VAR_GLOBAL   // PLC tag table "RIO_6"
   "Tank 6P GTT Isolation Valve Feedback - Opened" AT %I60.0 : Bool;   // CV422-6P
   "Tank 6P GTT Isolation Valve Feedback - Closed" AT %I60.1 : Bool;   // CV422-6P
   "Tank 6P Tank Vent Valve 1 Feedback - Opened" AT %I60.2 : Bool;   // CV441-6PA
   "Tank 6P Tank Vent Valve 1 Feedback - Closed" AT %I60.3 : Bool;   // CV441-6PA
   "Tank 6P Tank Vent Valve 2 Feedback - Opened" AT %I60.4 : Bool;   // CV441-6PB
   "Tank 6P Tank Vent Valve 2 Feedback - Closed" AT %I60.5 : Bool;   // CV441-6PB
   "RIO6_SPR_DI_60_6" AT %I60.6 : Bool;   // Spare input
   "RIO6_SPR_DI_60_7" AT %I60.7 : Bool;   // Spare input
   "Tank 6S GTT Isolation Valve Feedback - Opened" AT %I63.0 : Bool;   // CV421-6S
   "Tank 6S GTT Isolation Valve Feedback - Closed" AT %I63.1 : Bool;   // CV421-6S
   "Tank 6S Tank Vent Valve 1 Feedback - Opened" AT %I63.2 : Bool;   // CV440-6SA
   "Tank 6S Tank Vent Valve 1 Feedback - Closed" AT %I63.3 : Bool;   // CV440-6SA
   "Tank 6S Tank Vent Valve 2 Feedback - Opened" AT %I63.4 : Bool;   // CV440-6SB
   "Tank 6S Tank Vent Valve 2 Feedback - Closed" AT %I63.5 : Bool;   // CV440-6SB
   "RIO6_SPR_DI_63_6" AT %I63.6 : Bool;   // Spare input
   "RIO6_SPR_DI_63_7" AT %I63.7 : Bool;   // Spare input
   "Tank 6P BWT Level High High Switch" AT %I66.0 : Bool;   // LS425-6P
   "RIO6 Tanks Pressure Switch Hi Hi" AT %I66.1 : Bool;   // PS436-6P/6S
   "Tank 6S BWT Level High High Switch" AT %I66.2 : Bool;   // LS422-6S
   "RIO6_SPR_DI_66_3" AT %I66.3 : Bool;   // Spare input
   "RIO6_SPR_DI_66_4" AT %I66.4 : Bool;   // Spare input
   "RIO6_SPR_DI_66_5" AT %I66.5 : Bool;   // Spare input
   "RIO6_SPR_DI_66_6" AT %I66.6 : Bool;   // Spare input
   "RIO6_SPR_DI_66_7" AT %I66.7 : Bool;   // Spare input
   "Tank 6P USD Flow Meter" AT %IW332 : Int;   // FIT418-6P
   "Tank 6P MBG Flow Meter" AT %IW334 : Int;   // FIT420-6P
   "Tank 6S USD Flow Meter" AT %IW336 : Int;   // FIT417-6S
   "Tank 6S MBG Flow Meter" AT %IW338 : Int;   // FIT419-6S
   "RIO6 Main Gas-To-Deck Pressure" AT %IW340 : Int;   // PT415
   "Tank 6P BWT Level" AT %IW342 : Int;   // LT422-6P
   "Tank 6S BWT Level" AT %IW344 : Int;   // LT421-6S
   "RIO6_SPR_AI_346" AT %IW346 : Int;   // Spare input
   "Tank 6P BWT ph" AT %IW348 : Int;   // 426-6P
   "Tank 6P BWT Temp" AT %IW350 : Int;   // 426-6P
   "Tank 6P BWT DO" AT %IW352 : Int;   // 428-6P
   "RIO6 Tanks Pressure" AT %IW354 : Int;   // PT424-6P/6S
   "Tank 6S BWT ph" AT %IW356 : Int;   // 425-6S
   "Tank 6S BWT Temp" AT %IW358 : Int;   // 425-6S
   "Tank 6S BWT DO" AT %IW360 : Int;   // 427-6S
   "RIO6_SPR_AI_362" AT %IW362 : Int;   // Spare input
   "Tank 6P Vent Valve 1" AT %Q20.0 : Bool;   // CV441-6PA
   "Tank 6P Vent Valve 2" AT %Q20.1 : Bool;   // CV441-6PB
   "Tank 6S Vent Valve 1" AT %Q20.2 : Bool;   // CV440-6SA
   "Tank 6S Vent Valve 2" AT %Q20.3 : Bool;   // CV440-6SB
END_VAR

VAR_GLOBAL   // PLC tag table "RIO_7"
   "APT GTT Isolation Valve Feedback - Opened" AT %I75.0 : Bool;   // CV422-APT
   "APT GTT Isolation Valve Feedback - Closed" AT %I75.1 : Bool;   // CV422-APT
   "APT Tank Vent Valve 1 Feedback - Opened" AT %I75.2 : Bool;   // CV441-APTA
   "APT Tank Vent Valve 1 Feedback - Closed" AT %I75.3 : Bool;   // CV441-APTA
   "APT Tank Vent Valve 2 Feedback - Opened" AT %I75.4 : Bool;   // CV441-APTB
   "APT Tank Vent Valve 2 Feedback - Closed" AT %I75.5 : Bool;   // CV441-APTB
   "RIO7_SPR_DI_175_6" AT %I75.6 : Bool;   // Spare input
   "RIO7_SPR_DI_175_7" AT %I75.7 : Bool;   // Spare input
   "APT BWT Level High High Switch" AT %I78.0 : Bool;   // LS425-APT
   "RIO7 Tank Pressure Switch Hi Hi" AT %I78.1 : Bool;   // PS436-APT
   "RIO7_SPR_DI_178_2" AT %I78.2 : Bool;   // Spare input
   "RIO7_SPR_DI_178_3" AT %I78.3 : Bool;   // Spare input
   "RIO7_SPR_DI_178_4" AT %I78.4 : Bool;   // Spare input
   "RIO7_SPR_DI_178_5" AT %I78.5 : Bool;   // Spare input
   "RIO7_SPR_DI_178_6" AT %I78.6 : Bool;   // Spare input
   "RIO7_SPR_DI_178_7" AT %I78.7 : Bool;   // Spare input
   "APT USD Flow Meter" AT %IW400 : Int;   // FIT418-APT
   "APT MBG Flow Meter" AT %IW402 : Int;   // FIT420-APT
   "RIO7 Confined Space O2 Monitor" AT %IW404 : Int;   // 600-TX-433
   "RIO7_SPR_AI_406" AT %IW406 : Int;   // Spare input
   "RIO7 Deck Main Pressure" AT %IW408 : Int;   // PT415
   "APT BWT Level" AT %IW410 : Int;   // LT422-APT
   "RIO7_SPR_AI_412" AT %IW412 : Int;   // Spare input
   "RIO7_SPR_AI_414" AT %IW414 : Int;   // Spare input
   "APT BWT ph" AT %IW416 : Int;   // 426-APT
   "APT BWT Temp" AT %IW418 : Int;   // 426-APT
   "APT BWT DO" AT %IW420 : Int;   // 428-APT
   "RIO7 Tank Pressure" AT %IW422 : Int;   // PT424-APT
   "APT Vent Valve 1" AT %Q26.0 : Bool;   // CV441-APTA
   "APT Vent Valve 2" AT %Q26.1 : Bool;   // CV441-APTB
   "RIO7_SPR_DQ_26_2" AT %Q26.2 : Bool;   // Spare output
   "600-TX-433 O2 Monitor Alarm" AT %Q26.3 : Bool;   // 600-TX-433 RIO7 Confined Space O2 Monitor
END_VAR

VAR_GLOBAL   // PLC tag table "WBT"
   "IN_Level_FPT" AT %IW1000 : Int;
   "IN_Level_WBT_1S" AT %IW1002 : Int;
   "IN_Level_WBT_1P" AT %IW1004 : Int;
   "IN_Level_WBT_2S" AT %IW1006 : Int;
   "IN_Level_WBT_2P" AT %IW1008 : Int;
   "IN_Level_WBT_3S" AT %IW1010 : Int;
   "IN_Level_WBT_3P" AT %IW1012 : Int;
   "IN_Level_WBT_4S" AT %IW1014 : Int;
   "IN_Level_WBT_4P" AT %IW1016 : Int;
   "IN_Level_WBT_5S" AT %IW1018 : Int;
   "IN_Level_WBT_5P" AT %IW1020 : Int;
   "IN_Level_WBT_6S" AT %IW1022 : Int;
   "IN_Level_WBT_6P" AT %IW1024 : Int;
   "IN_Level_APT" AT %IW1026 : Int;
END_VAR

// folder: Alarms & Sensors

TYPE "ANALOG_SENSOR_LIMITS"
   STRUCT
      Minimum : Real;   // Minimum sensor limit
      Maximum : Real;   // Maximum sensor limit
   END_STRUCT;
END_TYPE

TYPE "ANALOG_SENSOR_SETPOINTS"
   STRUCT
      LowLow : Real;   // Setpoint for LowLow
      Low : Real;   // Setpoint for Low
      High : Real;   // Setpoint for High
      HighHigh : Real;   // Setpoint for HighHigh
   END_STRUCT;
END_TYPE

TYPE "ANALOG_SENSOR_4_ALARMS"
   STRUCT
      Healthy : Bool;   // This sensor is healthy (no alarms)
      LowLow : Bool;   // Sensor reporting under LowLow setpoint
      Low : Bool;   // Sensor reporting under Low setpoint but above LowLow
      High : Bool;   // Sensor reporting above High setpoint but below HighHigh setpoint
      HighHigh : Bool;   // Sensor reporting above HighHigh setpoint
   END_STRUCT;
END_TYPE

TYPE "ANALOG_SENSOR_2_ALARMS"
   STRUCT
      Healthy : Bool;   // This sensor is healthy (no alarms)
      Low : Bool;   // Sensor reporting under Low setpoint
      High : Bool;   // Sensor reporting above High setpoint
   END_STRUCT;
END_TYPE

TYPE "VALVE_STATES"
   STRUCT
      Open : Bool;   // Valve is open {OPEN=True, CLSD=False}
      Closed : Bool;   // Valve is closed {OPEN=False, CLSD=True}
      Moving : Bool;   // Valve is moving {OPEN=False, CLSD=False}
      Fault : Bool;   // Valve is in error {OPEN=True, CLSD=True}
   END_STRUCT;
END_TYPE

TYPE "DIGITAL_SENSOR_ALARMS"
   STRUCT
      Healthy : Bool;   // Is this sensor Healthy?
      UnhealthyAlarm : Bool;   // Has an alarm been raised? (Low/High depending on Sensor type)
   END_STRUCT;
END_TYPE

// folder: Auto BWT Sequencing

TYPE "TANK_DATA"
   STRUCT
      TankID : Int := 0;   // Tank ID of this object.
      TankState : Int := 0;   // Describes the state which this tank is currently in. Allows for differentation between system state and tank sub state due to treatment groups architecture allowing multuple states at one time.
      Active : Bool := false;   // Is this tank active (data populated from Adj. Consts)
      AllocatedTreatmentGroup : Int := 0;   // Describes which treatment group this tank is allocated to. This data is hard-coded in any instantiation of this data type.
      XeOx_Complete : Bool := false;   // Reports ReOx/DeOx completion (same variable reused for simplification of code as ReOx and DeOx are mutually exclusive).
      Timer_Complete : Bool := false;   // Reports MId-Dwell/Post-Dwell timer completion (same variable reused for simplification of code as Mid-Dwell and Post-Dwell are mutually exclusive).
   END_STRUCT;
END_TYPE

TYPE "SYSTEM_STATES"
   STRUCT
      System : Int;   // Describes the overall system state.
      DeOx : Int;   // Describes the DeOx sub-state in action.
      ReOx : Int;   // Describes the ReOx sub-state in action.
      Complete : Int;   // Describes the Completion sub-state in action.
      TreatmentGroup : Int;   // Identifies which TreatmentGroup is currently being actioned. This is re-used in ReOx and DeOx modes of operation as they are mutually exclusive.
   END_STRUCT;
END_TYPE

TYPE "ALARM_DEMAND_RTN"
   STRUCT
      Demand_Complete : Bool;   // Has the demand been completed? {T:Demand is complete;F:Demand is not yet complete, timer has not timed out}
      Alarm_Active : Bool;   // Has an alarm been raised? {T:Timeout has ocurred valve failed to actuate;F:No active alarm valve is still actuating}
   END_STRUCT;
END_TYPE

TYPE "GTT_EXCLUSIVITY"
   STRUCT
      Tank_Exclusivity : Bool;   // Is a GTT Valve currently in operation (openning or closing)
      TankID_InOperation : Int;   // The Tank ID number which is currently in transition
   END_STRUCT;
END_TYPE

TYPE "HMI_MESSAGE"
   STRUCT
      Active : Bool;   // Should the alert be displayed?
      Message : String;   // What alert should be displayed?
   END_STRUCT;
END_TYPE

TYPE "VALVE_PVVX_IN"
   STRUCT
      PVVx_Actuate : Array[1..14] of Bool;
      PVVA_ValveDemands : Array[1..14] of Bool;
      PVVB_ValveDemands : Array[1..14] of Bool;
   END_STRUCT;
END_TYPE

TYPE "VALVE_GTT_IN"
   STRUCT
      GTT_Actuate : Array[1..14] of Bool;
      GTT_ValveDemands : Array[1..14] of Bool;
   END_STRUCT;
END_TYPE

TYPE "VALVE_PVVX_OUT"
   STRUCT
      PVVA_DemandsCompleted : Array[1..14] of Bool;
      PVVA_Alarms : Array[1..14] of Bool;
      PVVB_DemandsCompleted : Array[1..14] of Bool;
      PVVB_Alarms : Array[1..14] of Bool;
   END_STRUCT;
END_TYPE

TYPE "VALVE_GTT_OUT"
   STRUCT
      GTT_DemandsCompleted : Array[1..14] of Bool;
      GTT_Alarms : Array[1..14] of Bool;
   END_STRUCT;
END_TYPE

// folder: Data Processing

TYPE "AI_DATA"
VERSION : 0.1
   STRUCT
      RAW_MIN : Int;   // Raw minimum value from AI card
      RAW_MAX : Int := 27648;   // Raw maximum value from AI card
      NORM : Real;   // Normalised real value
      ENG_MIN : Real;   // Engineering units minimum value
      ENG_MAX : Real := 100.0;   // Engineering units maximum value
   END_STRUCT;
END_TYPE

TYPE "AQ_DATA"
VERSION : 0.1
   STRUCT
      ENG_MIN : Real;   // Engineering units minimum value
      ENG_MAX : Real := 100.0;   // Engineering units maximum value
      NORM : Real;   // Normalised real value
      RAW_MIN : Int;   // Raw minimum value from AQ card
      RAW_MAX : Int := 27648;   // Raw maximum value from AQ card
   END_STRUCT;
END_TYPE

TYPE "TANK_IP_DATA"
VERSION : 0.1
   STRUCT
      O2_MONITOR : Real;   // Space monitor, 600-Tx-433
      DECK_IG_PRESS : Real;   // Deck main IG pressure, PT-415
      TANKS_PRESS : Real;   // Tank group pressure, PT-424
      TANKS_PRESS_HIHI : Bool;   // Tank group pressure, PS-436
      TANK_GROUP_SPARE_DI_2 : Bool;   // Spare input
      TANK_GROUP_SPARE_DI_3 : Bool;   // Spare input
      TANK_GROUP_SPARE_DI_4 : Bool;   // Spare input
      TANK_GROUP_SPARE_DI_5 : Bool;   // Spare input
      TANK_GROUP_SPARE_DI_6 : Bool;   // Spare input
      TANK_GROUP_SPARE_DI_7 : Bool;   // Spare input
      GTT_ISOL_VALVE_OPEN : Bool;   // Gas to tank isolation valve feedback, CV-422
      GTT_ISOL_VALVE_CLSD : Bool;   // Gas to tank isolation valve feedback, CV-422
      TANK_VENT_A_OPEN : Bool;   // Tank vent valve feedback, CV-441-A
      TANK_VENT_A_CLSD : Bool;   // Tank vent valve feedback, CV-441-A
      TANK_VENT_B_OPEN : Bool;   // Tank vent valve feedback, CV-441-B
      TANK_VENT_B_CLSD : Bool;   // Tank vent valve feedback, CV-441-B
      BWT_LEVEL_HIHI : Bool;   // Tank water level, LS-425
      TANK_ALARM : Bool;   // Tank Alarm
      SPARE_DI_7 : Bool;   // Spare input
      USD_FLOW : Real;   // FIT-418
      "USD FLOW  N" : Real;
      MBG_FLOW : Real;   // FIT-420
      "MBG_FLOW N" : Real;
      BWT_LEVEL : Real;   // LT-422
      BWT_PH : Real;   // Ph 426
      BWT_TEMP : Real;   // Temperature 426
      BWT_DO : Real;   // Disolved oxygen 428
      SPARE_AI_1 : Real;   // Spare input
      SPARE_AI_2 : Real;   // Spare input
      SPARE_AI_3 : Real;   // Spare input
      USD_FLOW_CNFG : "AI_DATA";   // Input processing configuration data
      MBG_FLOW_CNFG : "AI_DATA";   // Input processing configuration data
      BWT_LEVEL_CNFG : "AI_DATA";   // Input processing configuration data
      BWT_PH_CNFG : "AI_DATA";   // Input processing configuration data
      BWT_TEMP_CNFG : "AI_DATA";   // Input processing configuration data
      BWT_DO_CNFG : "AI_DATA";   // Input processing configuration data
      SPARE_AI_1_CNFG : "AI_DATA";   // Input processing configuration data
      SPARE_AI_2_CNFG : "AI_DATA";   // Input processing configuration data
      SPARE_AI_3_CNFG : "AI_DATA";   // Input processing configuration data
      O2_MONITOR_CNFG : "AI_DATA";   // Input processing configuration data
      DECK_IG_PRESS_CNFG : "AI_DATA";   // Input processing configuration data
      TANKS_PRESS_CNFG : "AI_DATA";   // Input processing configuration data
   END_STRUCT;
   // BWT_DO_CNFG.ENG_MAX := 20.0;
   // USD_FLOW_CNFG.ENG_MAX := 55.0;
   // MBG_FLOW_CNFG.ENG_MAX := 23.0;
   // BWT_PH_CNFG.ENG_MAX := 12.0;
   // BWT_PH_CNFG.ENG_MIN := 2.0;
   // BWT_TEMP_CNFG.ENG_MIN := -15.0;
   // BWT_TEMP_CNFG.ENG_MAX := 80.0;
   // O2_MONITOR_CNFG.ENG_MAX := 15.0;
   // DECK_IG_PRESS_CNFG.ENG_MAX := 10.0;
   // TANKS_PRESS_CNFG.ENG_MIN := -200.0;
   // TANKS_PRESS_CNFG.ENG_MAX := 200.0;
END_TYPE

TYPE "1T_IP_DATA"
VERSION : 0.1
   STRUCT
      FIRST_TANK : "TANK_IP_DATA";
   END_STRUCT;
END_TYPE

TYPE "2T_IP_DATA"
VERSION : 0.1
   STRUCT
      FIRST_TANK : "TANK_IP_DATA";
      SECOND_TANK : "TANK_IP_DATA";
   END_STRUCT;
END_TYPE

TYPE "3T_IP_DATA"
VERSION : 0.1
   STRUCT
      FIRST_TANK : "TANK_IP_DATA";
      SECOND_TANK : "TANK_IP_DATA";
      THIRD_TANK : "TANK_IP_DATA";
   END_STRUCT;
END_TYPE

// folder: 10 - 19 IO & Processing

DATA_BLOCK "10_DI_DATA"   // DB10
TITLE = Digital Input Data
{ S7_Optimized_Access := 'TRUE' }
AUTHOR : JRS
VERSION : 0.1
// Processed data for code use
   VAR
      R3_SPR_DI_136_0 : Bool;   // Spare input
      R3_SPR_DI_136_1 : Bool;   // Spare input
      "FS_332 FLW_OK" : Bool;   // Cooling seawater flow switch
      CV358_OPN : Bool;   // FW Fill valve feedback open
      CV358_CLSD : Bool;   // FW Fill valve feedback closed
      FS_350_FLW_OK : Bool;   // Fresh water cooling flow switch
      CV341_OPN : Bool;   // GCU Drain valve feedback open
      CV341_CLSD : Bool;   // GCU Drain valve feedback closed
      CV406_OPN : Bool;   // Gas to deck valve feedback open
      CV406_CLSD : Bool;   // Gas to deck valve feedback closed
      CV407_OPN : Bool;   // Gas block valve 1 feedback open
      CV407_CLSD : Bool;   // Gas block valve 1 feedback closed
      CV411_OPN : Bool;   // Gas block valve 2 feedback open
      CV411_CLSD : Bool;   // Gas block valve 2 feedback closed
      CV409_OPN : Bool;   // Gas bleed valve feedback open
      CV409_CLSD : Bool;   // Gas bleed valve feedback closed
      CV441_OPN : Bool;   // Ambient air valve feedback open
      CV441_CLSD : Bool;   // Ambient air valve feedback closed
      LS_303_LO : Bool;   // GCU Low level switch
      P_304_ENBLD : Bool;   // GCU Booster pump enabled
      PB_10S1 : Bool;   // GCU Local PB - Start
      PB_10S2 : Bool;   // GCU Local PB - Stop
      EPB_8S1 : Bool;   // E-Stop Pressed @ BWT CP
      P_303_ENBLD : Bool;   // GCU Recirculation pump enabled
      E_400_STPD : Bool;   // Process gas compressor running/stopped
      E_400_SHTDN : Bool;   // Process gas compressor tripped/shutdown
      P_303_OK : Bool;   // GCU Recirculation pump healthy
      "5T1_PWR_OK" : Bool;   // 5T1 Power healthy
      "6Q6_PWR_OK" : Bool;   // Panel vent power healthy
      P_304_OK : Bool;   // GCU Booster pump healthy
      E_400_RUN : Bool;   // PGC Running loaded/on-line
      E_400_NOK : Bool;   // PGC Alarm/warning
   END_VAR
BEGIN
END_DATA_BLOCK

DATA_BLOCK "12_AI_Data"   // DB12
TITLE = Analogue Input Data
{ S7_Optimized_Access := 'TRUE' }
AUTHOR : JRS
VERSION : 0.1
// Processed data for code use
   VAR
      LIT_304_SCALED : Real;   // GCU Level
      R3_SPR_AI_802_SCALED : Real;   // BWT Control panel temperature
      TIT_408_SCALED : Real;   // Fresh water cooling temperature
      TIT_406_SCALED : Real;   // Gas to deck (Outlet) temperature
      CV_405_SCALED : Real;   // Gas To deck vent valve feedback
      PIT_416_SCALED : Real;   // Gas to deck pressure
      PIT_358_SCALED : Real;   // Fresh water inlet pressure
      PIT_348_SCALED : Real;   // GCU Cooling seawater pressure
      PIT_353_SCALED : Real;   // Recirculation fresh water pressure
      E_400_PT002_SCALED : Real;   // PGC Discharge (outlet) pressure
      E_400_TE002_SCALED : Real;   // PGC Discharge (outlet) temperature
      SL_400_SCALED : Real;   // Ballast water salinity
      R3_SPR_AI_824_SCALED : Real;   // Spare input
      R3_SPR_AI_826_SCALED : Real;   // Spare input
      R3_SPR_AI_828_SCALED : Real;   // Spare input
      R3_SPR_AI_830_SCALED : Real;   // Spare input
      IW_800 : "AI_DATA";   // IW800 - GCU Level (LIT-304)
      IW_802 : "AI_DATA";   // IW802 - BWT Control Panel Temperature (PT-100)
      IW_804 : "AI_DATA";   // IW804 - Fresh Water Cooling Temperature (TIT-408)
      IW_806 : "AI_DATA";   // IW806 - Gas to Deck Outlet Temperature (TIT-406)
      IW_808 : "AI_DATA";   // IW808 - Gas to Deck Vent Valve Feedback (CV-405)
      IW_810 : "AI_DATA";   // PIT416
      IW_812 : "AI_DATA";   // PIT358
      IW_814 : "AI_DATA";   // PIT348
      IW_816 : "AI_DATA";   // PIT353
      IW_818 : "AI_DATA";   // E400-PT002
      IW_820 : "AI_DATA";   // E400-TT002
      IW_822 : "AI_DATA";   // SL-400
      IW_824 : "AI_DATA";   // Spare input
      IW_826 : "AI_DATA";   // Spare input
      IW_828 : "AI_DATA";   // Spare input
      IW_830 : "AI_DATA";   // Spare input
   END_VAR
BEGIN
   IW_806.ENG_MIN := 0.0;
   IW_806.ENG_MAX := 150.0;
   IW_804.ENG_MIN := 0.0;
   IW_804.ENG_MAX := 150.0;
   IW_816.ENG_MAX := 10.0;
   IW_810.ENG_MAX := 10.0;
   IW_812.ENG_MAX := 10.0;
   IW_814.ENG_MAX := 10.0;
   IW_818.ENG_MAX := 6.0;
   IW_820.ENG_MAX := 300.0;
END_DATA_BLOCK

DATA_BLOCK "14_DQ_DATA"   // DB14
TITLE = Digital Output Data
{ S7_Optimized_Access := 'TRUE' }
AUTHOR : JRS
VERSION : 0.1
// Processed data for output via physical connection
   VAR
      CV_358 : Bool;   // Fresh water fill valve control
      CV_341 : Bool;   // Waste water drain valve control
      CV_407 : Bool;   // Block valve 1 control
      CV_409 : Bool;   // Bleed valve control
      CV_411 : Bool;   // Block valve 2 control
      CV_441 : Bool;   // Ambient air valve control
      CV_406 : Bool;   // Main gas to deck valve control
      E_400_RUN : Bool;   // Start process gas compressor
      P_303 : Bool;   // GCU Recirculation pump control
      P_304 : Bool;   // GCU Booster pump control
      "13P1" : Bool;   // GCU Warning alarm
      "13P2" : Bool;   // GCU Shutdown alarm
      "13P3" : Bool;   // GCU Running
      "13P4" : Bool;   // Ballast water tank level HIHI
      "13P5" : Bool;   // GCU Alarm buzzer
      E_400_STP : Bool;   // Stop process gas compressor
      CV_422_FPT : Bool;   // Pilot for GTT FPT Valve
      CV_422_1P : Bool;   // Pilot for GTT 1 Port valve
      CV_421_1S : Bool;   // Pilot for GTT 1 Starboard valve
      CV_422_2P : Bool;   // Pilot for GTT 2 Port valve
      CV_421_2S : Bool;   // Pilot for GTT 2 Starboard valve
      CV_422_3P : Bool;   // Pilot for GTT 3 Port valve
      CV_421_3S : Bool;   // Pilot for GTT 3 Starboard valve
      R3_SPR_DQ_138_7 : Bool;   // Spare output
      CV_422_4P : Bool;   // Pilot for GTT 4 Port valve
      CV_421_4S : Bool;   // Pilot for GTT 4 Starboard valve
      CV_422_5P : Bool;   // Pilot for GTT 5 Port valve
      CV_421_5S : Bool;   // Pilot for GTT 5 Starboard valve
      CV_422_6P : Bool;   // Pilot for GTT 6 Port valve
      CV_421_6S : Bool;   // Pilot for GTT 6 Starboard valve
      CV_422_APT : Bool;   // Pilot for GTT APT Port valve
      R3_SPR_DQ_139_7 : Bool;   // Spare output
   END_VAR
BEGIN
END_DATA_BLOCK

DATA_BLOCK "16_AQ_Data"   // DB16
TITLE = Analogue Output Data
{ S7_Optimized_Access := 'TRUE' }
AUTHOR : JRS
VERSION : 0.1
// Processed data for output via physical connection
   VAR RETAIN
      CV405_CNTRL : Real;   // Gas vent position control
   END_VAR
   VAR
      R3_SPR_AQ_802 : Real;   // Spare output
      R3_SPR_AQ_804 : Real;   // Spare output
      R3_SPR_AQ_806 : Real;   // Spare output
      QW_800 : "AQ_DATA";   // Output word data, edit calibration here
      QW_802 : "AQ_DATA";   // Output word data, edit calibration here
      QW_804 : "AQ_DATA";   // Output word data, edit calibration here
      QW_806 : "AQ_DATA";   // Output word data, edit calibration here
   END_VAR
BEGIN
END_DATA_BLOCK

DATA_BLOCK "19_AUTO_CMNDS_Data"   // DB19
TITLE = Automatic Commands Data
{ S7_Optimized_Access := 'TRUE' }
AUTHOR : JRS
VERSION : 0.1
// Defined data for use prior to output processing
   VAR
      PIT416_CMND_Target : Real := 0.0;   // PIT416 Commanded target (bar g)
      LIT304_CMND_Target : Real := 61.0;   // LIT304 Commanded target (%) [GEN-19]
      LIT304_CMND_Target_Low : Real;
      LIT304_CMND_LowLow : Real := 33.0;   // LIT304 Commanded low low setpoint (%) [GEN-19]
      LIT304_CMND_Low : Real := 44.0;   // LIT304 Commanded low set point (%) [GEN-19]
      LIT304_CMND_High : Real := 78.0;   // LIT304 Commanded high setpoint (%) [GEN-19]
      LIT304_CMND_HighHigh : Real := 89.0;   // LIT304 Commanded high high setpoint (%)
      PIT353_CMND_LowLow : Real := 1.0;   // PIT353 Commanded low low setpoint (bar g)
      PIT353_CMND_Low : Real := 1.5;   // PIT353 Commanded low setpoint (bar g)
      PIT353_CMND_High : Real := 3.5;   // PIT353 Commanded high setpoint (bar g)
      PIT353_CMND_HighHigh : Real := 4.0;   // PIT353 Commanded high high setpoint (bar g)
      PIT358_CMND_LowLow : Real := 1.0;   // PIT358 Commanded low low setpoint (bar g)
      PIT358_CMND_Low : Real := 1.5;   // PIT358 Commanded low setpoint (bar g)
      PIT358_CMND_High : Real := 3.5;   // PIT358 Commanded high setpoint (bar g)
      PIT358_CMND_HighHigh : Real := 4.0;   // PIT358 Commanded high high setpoint (bar g)
      CV405_PID_MDLTG : Bool;   // 1 = Modulating, 0 = Not
      CV401_CLS_FLAG : Bool;   // 1 = Close, 0 = Not
      CV441_OPN_FLG : Bool;   // 1 = Open, 0 = Not
      WRNG_PLS : Bool;   // Pulse bit
      ALRM_PLS : Bool;   // Pulse bit
      BTCS_ACTV : Bool;   // 1 = Active, 0 = Not
      ACTV_PLS : Bool;   // Pulse bit
      "Purge Rqst Simulate" : Bool;
   END_VAR
BEGIN
END_DATA_BLOCK

DATA_BLOCK "PGC Flush_DB"   // DB23
{ S7_Optimized_Access := 'TRUE' }
VERSION : 0.1
// stored: InstanceOfName PGC Flush
"PGC Flush"
BEGIN
END_DATA_BLOCK

// folder: 100 - 199 Automatic Sequencing

DATA_BLOCK "100_GCU_AUTO_SEQ_DB"   // DB100
TITLE = GCU Auto Sequence Instance DB
{ S7_Optimized_Access := 'TRUE' }
AUTHOR : JRS
VERSION : 0.1
// Data required for FB
// stored: InstanceOfName 100_GCU_AUTO_SEQ
"100_GCU_AUTO_SEQ"
BEGIN
END_DATA_BLOCK

DATA_BLOCK "Setpoint Override_DB"   // DB104
{ S7_Optimized_Access := 'TRUE' }
VERSION : 0.1
// stored: InstanceOfName Setpoint Override
"Setpoint Override"
BEGIN
END_DATA_BLOCK

DATA_BLOCK "RAMP_DB"   // DB105
{ S7_Optimized_Access := 'TRUE' }
VERSION : 0.1
// stored: InstanceOfName RAMP
"RAMP"
BEGIN
END_DATA_BLOCK

DATA_BLOCK "Tank Change"   // DB106
{ S7_Optimized_Access := 'TRUE' }
VERSION : 0.1
// stored: InstanceOfName Binary Imputs ADD
"Binary Imputs ADD"
BEGIN
END_DATA_BLOCK

DATA_BLOCK "108_GCU_TNK_REFILL_SEQ_DB"   // DB108
{ S7_Optimized_Access := 'TRUE' }
AUTHOR : JRS
VERSION : 0.1
// stored: InstanceOfName 108_GCU_TNK_REFILL_SEQ
"108_GCU_TNK_REFILL_SEQ"
BEGIN
END_DATA_BLOCK

DATA_BLOCK "109_TRGT_RAMP_CNTRL_DB"   // DB109
{ S7_Optimized_Access := 'TRUE' }
AUTHOR : JRS
VERSION : 0.1
// stored: InstanceOfName 109_TRGT_RAMP_CNTRL
"109_TRGT_RAMP_CNTRL"
BEGIN
END_DATA_BLOCK

DATA_BLOCK "110_GCU_TNK_FLUSH_SEQ_DB"   // DB110
{ S7_Optimized_Access := 'TRUE' }
AUTHOR : JRS
VERSION : 0.1
// stored: InstanceOfName 110_GCU_TNK_FLUSH_SEQ
"110_GCU_TNK_FLUSH_SEQ"
BEGIN
END_DATA_BLOCK

DATA_BLOCK "140_PGC_HRS_RUN_DB"   // DB140
{ S7_Optimized_Access := 'TRUE' }
AUTHOR : JRS
VERSION : 0.1
// stored: InstanceOfName 140_PGC_HRS_RUN
"140_PGC_HRS_RUN"
BEGIN
END_DATA_BLOCK

DATA_BLOCK "141_P303_HRS_RUN_DB"   // DB141
{ S7_Optimized_Access := 'TRUE' }
AUTHOR : JRS
VERSION : 0.1
// stored: InstanceOfName 141_P303_HRS_RUN
"141_P303_HRS_RUN"
BEGIN
END_DATA_BLOCK

DATA_BLOCK "142_P304_HRS_RUN_DB"   // DB142
{ S7_Optimized_Access := 'TRUE' }
AUTHOR : JRS
VERSION : 0.1
// stored: InstanceOfName 142_P304_HRS_RUN
"142_P304_HRS_RUN"
BEGIN
END_DATA_BLOCK

DATA_BLOCK "150_GCU_LCL_CNTRL_DB"   // DB150
TITLE = GCU Local Control Data
{ S7_Optimized_Access := 'TRUE' }
AUTHOR : JRS
VERSION : 0.1
// Data area for local and automatic control of the GCU
   VAR
      LCL_CNTRL_ACTV : Bool := false;   // 1 = Local control active, 0 = Not (Tank System)
      SYS_OK_FOR_LCL : Bool := false;   // 1 = System ok for local control, 0 = Not
      STRT_AIR : Bool := false;   // 1 = Start with air command from HMI, 0 = Not
      STRT_IG : Bool := false;   // 1 = Start with IG command from HMI, 0 = Not
      STOP : Bool := false;   // 1 = Stop command
      RUN_WITH_AIR : Bool := false;   // 1 = Running with air, 0 = Not
      RUN_WITH_IG : Bool := false;   // 1 = Running with IG, 0 = Not
      TEST_BIT_1 : Bool := false;   // 1 = Test active, 0 = Not (commissioning bit)
      OPN_ACTV_GTT_VLVS : Bool;   // 1 = Open Active Valves, 0 = Not
      PLS_1 : Bool;   // Pulse bit
      PLS_2 : Bool;
   END_VAR
BEGIN
END_DATA_BLOCK

// folder: 1000 - 1999 BWT System Control/1090 - 1099 HMI Handling

DATA_BLOCK "721_VLV_CHK_DB"   // DB721
{ S7_Optimized_Access := 'TRUE' }
AUTHOR : JRS
VERSION : 0.1
// stored: InstanceOfName 501_VLV_CHK
"501_VLV_CHK"
BEGIN
END_DATA_BLOCK

DATA_BLOCK "1090_HMI_IP_FLAGS"   // DB1090
{ S7_Optimized_Access := 'TRUE' }
VERSION : 0.1
   VAR
      StartTreatment : Bool;   // Flag to BWTS to start treatment (BMWS-068)
      StopTreatment : Bool;   // Flag to BWTS to stop treatment
      BWTOperatingMode : Bool;   // True=Automatic BWTS, False=Manual Control
      BWTWithCB : Bool;
      ShipsLevelSensors : Bool;   // What type of sensors are in use on this system - True=Ship supplied, False=CHM supplied.
      PressVacuumValves : Bool;   // Is this system setup with pressure vacuum valves?
      ManualDemand_VentA : Array[1..14] of Bool;
      ManualDemand_VentB : Array[1..14] of Bool;
      ManualDemand_GTT : Array[1..14] of Bool;
   END_VAR
BEGIN
END_DATA_BLOCK

DATA_BLOCK "1092_HMI_OP_FLAGS"   // DB1092
{ S7_Optimized_Access := 'TRUE' }
VERSION : 0.1
   VAR
      HMI_Warnings : "HMI_MESSAGE";   // StartIGGWarnings / ReOxygenationWarning
      PIT415_Alarms : "ANALOG_SENSOR_4_ALARMS";   // Alarm (BWMS-020)
      "600CV407_Alarms" : "VALVE_STATES";   // Alarm (BWMS-020)
      "600CV409_Alarms" : "VALVE_STATES";   // Alarm (BWMS-020)
      "600CV411_Alarms" : "VALVE_STATES";   // Alarm (BWMS-020)
      TX430_Low_Alarm : Bool;   // Alarm (BWMS-020)
      TX425_426_pH_Alarms : Array[1..14] of "ANALOG_SENSOR_2_ALARMS";   // Alarm (BWMS-021)
      TX427_428_DO_Alarms : Array[1..14] of "ANALOG_SENSOR_2_ALARMS";   // Alarm (BWMS-021)
      FIT417_418_USDFlow_Alarms : Array[1..14] of "ANALOG_SENSOR_4_ALARMS";   // Alarm (BWMS-021)
      FIT419_420_MBGFlow_Alarms : Array[1..14] of "ANALOG_SENSOR_4_ALARMS";   // Alarm (BWMS-021)
      LT421_422_BWTLevel_Alarms : Array[1..14] of "ANALOG_SENSOR_2_ALARMS";   // Alarm (BWMS-021)
      LS425_442_LevelSwitch_HighHigh_Alarm : Array[1..14] of "DIGITAL_SENSOR_ALARMS";   // Alarm (BWMS-021)
      CV421_422_InletValve_Alarms : Array[1..14] of "VALVE_STATES";   // Alarm (BWMS-021)
      CV427_428_PVVA_Alarms : Array[1..14] of "VALVE_STATES";   // Alarm (BWMS-021)
      CV429_430_PVVB_Alarms : Array[1..14] of "VALVE_STATES";   // Alarm (BWMS-021)
      PT424_Alarms : Array[1..7] of "ANALOG_SENSOR_4_ALARMS";   // Alarm (BWMS-022)
      PS436_HighHigh_Alarm : Array[1..7] of "DIGITAL_SENSOR_ALARMS";   // Alarm (BWMS-022)
      NoTanksActive : Bool := false;   // Flag to show alert on HMI if no tanks are active (BMWS-065)
      VoyageLessThanTreatmentTime : Bool := false;   // Flag to show alert on HMI if Voyage time is less than the treatment time (BMWS-067)
      DeckSupplyOk : Bool := false;   // Flag when deck supply is OK (BMWS-083)
      StartButtonEnabled : Bool;   // Flag to HMI to dictate if start button should be enabled
   END_VAR
BEGIN
   HMI_Warnings.Active := false;
END_DATA_BLOCK

DATA_BLOCK "1094_ANALOGUE_SENSOR_SETPOINTS"   // DB1094
{ S7_Optimized_Access := 'TRUE' }
VERSION : 0.1
   VAR
      FIT417_418 : Array[1..14] of "ANALOG_SENSOR_SETPOINTS";   // Setpoints for FIT417, FIT418
      FIT419_420 : Array[1..14] of "ANALOG_SENSOR_SETPOINTS";   // Setpoints for FIT419, FIT420
      LT421_422 : "ANALOG_SENSOR_SETPOINTS";   // Setpoints for LT421, LT422
      PIT415 : "ANALOG_SENSOR_SETPOINTS";   // Setpoints for PIT415
      PT424 : "ANALOG_SENSOR_SETPOINTS";   // Setpoints for PT424
      TX425_426 : "ANALOG_SENSOR_SETPOINTS";   // Setpoints for TX425, TX426
      TX427_428_DEOX : "ANALOG_SENSOR_SETPOINTS";   // Setpoints for TX427, TX428 during DeOx
      TX427_428_REOX : "ANALOG_SENSOR_SETPOINTS";   // Setpoints for TX427, TX428 during ReOx
      TX430 : "ANALOG_SENSOR_SETPOINTS";   // Setpoints for TX430 (aka SL400)
   END_VAR
BEGIN
   LT421_422.Low := 90.0;   // %
   LT421_422.High := 98.0;   // %
   PIT415.LowLow := 2.8;   // bar(g)
   PIT415.Low := 3.0;   // bar(g)
   PIT415.High := 4.5;   // bar(g)
   PIT415.HighHigh := 4.8;   // bar(g)
   PT424.LowLow := -0.07;   // bar(g)
   PT424.Low := -0.05;   // bar(g)
   PT424.High := 0.08;   // bar(g)
   PT424.HighHigh := 0.09;   // bar(g)
   TX427_428_DEOX.Low := 0.2;   // mg/L
   TX427_428_DEOX.High := 12.0;   // mg/L
   TX427_428_REOX.Low := 0.2;   // mg/L
   TX427_428_REOX.High := 12.0;   // mg/L
   TX425_426.Low := 5.0;   // pH
   TX425_426.High := 9.5;   // pH
   TX430.High := 40.0;
   TX430.HighHigh := 40.0;
   TX430.Low := 0.1;
   TX430.LowLow := 0.1;
END_DATA_BLOCK

DATA_BLOCK "1096_ADJUSTABLE_CONSTANTS"   // DB1096
{ S7_Optimized_Access := 'TRUE' }
VERSION : 0.1
   VAR
      "600CV407Open_Time" : LTime := LT#30s;   // Time
      "600CV407Close_Time" : LTime := LT#30s;   // Time
      "600CV409Open_Time" : LTime := LT#30s;   // Time
      "600CV409Close_time" : LTime := LT#30s;   // Time
      "600CV411Open_Time" : LTime := LT#30s;   // Time
      "600CV411Close_time" : LTime := LT#30s;   // Time
      BWTInletValveOpen_Time : LTime := LT#30s;   // Time
      BWTInletValveClose_Time : LTime := LT#30s;   // Time
      PVVOpen_Time : LTime := LT#30s;   // Time
      PVVClose_Time : LTime := LT#30s;   // Time
      PIT415Delay_Time : LTime := LT#30s;   // Time
      TX430LowSP : Real := 0.1;   // % low setpoint
      TankIDDeselectBWT : Array[1..14] of Bool;   // allow de-selection of tank.
      TankIDActive : Array[1..14] of Bool;   // is the Tank active?
      VoyageTime : LTime;   // Time in hours
   END_VAR
BEGIN
   TankIDActive[1] := true;
   TankIDActive[2] := true;
   TankIDActive[3] := true;
   TankIDActive[4] := true;
   TankIDActive[5] := true;
   TankIDActive[6] := true;
   TankIDActive[7] := true;
   TankIDActive[8] := true;
   TankIDActive[9] := true;
   TankIDActive[10] := true;
   TankIDActive[11] := true;
   TankIDActive[12] := true;
   TankIDActive[13] := true;
   TankIDActive[14] := true;
END_DATA_BLOCK

DATA_BLOCK "1098_ANALOGUE_SENSOR_LIMITS"   // DB1098
{ S7_Optimized_Access := 'TRUE' }
VERSION : 0.1
   VAR
      FIT417_418 : Array[1..14] of "ANALOG_SENSOR_LIMITS";   // Sensor Limits for FIT417, FIT418
      FIT419_420 : Array[1..14] of "ANALOG_SENSOR_LIMITS";   // Sensor Limits for FIT419, FIT420
      LT421_422 : "ANALOG_SENSOR_LIMITS";   // Sensor Limits for LT421, LT422
      PIT415 : "ANALOG_SENSOR_LIMITS";   // Sensor Limits for PIT415
      PT424 : "ANALOG_SENSOR_LIMITS";   // Sensor Limits for PT424
      TX425_426 : "ANALOG_SENSOR_LIMITS";   // Sensor Limits for TX425, TX426
      TX427_428 : "ANALOG_SENSOR_LIMITS";   // Sensor Limits for TX427, TX428
      TX430 : "ANALOG_SENSOR_LIMITS";   // Sensor Limits for TX430
   END_VAR
BEGIN
   PIT415.Maximum := 10.0;   // bar(g)
   PIT415.Minimum := 0.0;   // bar(g)
   LT421_422.Maximum := 98.0;   // %
   LT421_422.Minimum := 90.0;   // %
   PT424.Minimum := -0.2;   // bar(g)
   PT424.Maximum := 0.2;   // bar(g)
   TX425_426.Minimum := 0.0;   // pH
   TX425_426.Maximum := 14.0;   // pH
   TX427_428.Minimum := 0.0;   // mg/L
   TX427_428.Maximum := 15.0;   // mg/L
   TX430.Minimum := 0.0;   // %
   TX430.Maximum := 40.0;   // %
   // FIT417_418.Minimum : Nm^3/hr
   // FIT417_418.Maximum : Nm^3/hr
   // FIT419_420.Minimum : Nm^3/hr
   // FIT419_420.Maximum : Nm^3/hr
END_DATA_BLOCK

// folder: 1000 - 1999 BWT System Control/1100 - 1104 BWTS Control

DATA_BLOCK "1100_BWTS_CONTROL_DB"   // DB1100
{ S7_Optimized_Access := 'TRUE' }
VERSION : 0.1
// stored: InstanceOfName 1100_BWTS_CONTROL
"1100_BWTS_CONTROL"
BEGIN
END_DATA_BLOCK

DATA_BLOCK "1101_MANUAL_CONTROL_DB"   // DB1101
{ S7_Optimized_Access := 'TRUE' }
VERSION : 0.1
// stored: InstanceOfName 1101_RIO_MANUAL_CONTROL
"1101_RIO_MANUAL_CONTROL"
BEGIN
END_DATA_BLOCK

// folder: 1000 - 1999 BWT System Control/1190 - 1199 Data

DATA_BLOCK "1190_FIXED_CONSTANTS"   // DB1190
{ S7_Optimized_Access := 'TRUE' }
VERSION : 0.1
   VAR
      IGGDemand : Bool := false;
      PreDwell_Time : LTime := LT#18h;   // Time
      DeOxMin_Time : LTime := LT#12h;   // Time
      DeOxAtLevel_Time : LTime := LT#2h;   // Time
      ReOxMin_Time : LTime := LT#6h;   // Time
      ReOxAtLevel_Time : LTime := LT#2h;   // Time
      MidDwell_Time : LTime := LT#60h;   // Time
      PostDwell_Time : LTime := LT#12h;   // Time
      DeOxTargetDOLevel : Real := 0.5;   // mg/L
      ReOxTargetpHLevel : Real := 6.5;   // pH
      MaxDOPause_Time : LTime;   // Time (TBC)
      NumberOfTreatmentGroups : Int := 5;
      NumberOfTanks : Int := 14;
   END_VAR
BEGIN
END_DATA_BLOCK

DATA_BLOCK "1191_SYSTEM_VARIABLES"   // DB1191
{ S7_Optimized_Access := 'TRUE' }
VERSION : 0.1
   VAR
      NumberOfActiveTanks : Int := 0;
      DeselectAndActiveTanksComplete : Bool := false;
      MidDwell_ElapsedTime : LTime;
      FromIGG_InertGasReady : Bool := false;   // IGG->BWTS flag (BWMS-027)
      FromIGG_IGGDemand : Bool;   // IGG->BWTS flag (BWMS-027)
      ToIGG_BWTOperatingMode : Int;   // BWTS->IGG flag (BWMS-028)
      ToIGG_BWTwithCB : Bool;   // BWTS->IGG flag (BWMS-028)
      ToIGG_LIT305In : Bool;   // BWTS->IGG flag (BWMS-028)
      ToIGG_P305EnabledIn : Bool;   // BWTS->IGG flag (BWMS-028)
      ToIGG_P305TrippedIn : Bool;   // BWTS->IGG flag (BWMS-028)
      StartIGGWarningsTime : LTime;
      TreatmentTime : LTime;
   END_VAR
BEGIN
END_DATA_BLOCK

// folder: 20 - 49 RIO & Processing

